   438: 'Spare_Fault_438', class No Acknowledgement, trigger "DB302_HMI_Faults_Carrier6_Faults_3" bit 5
   439: 'Spare_Fault_439', class No Acknowledgement, trigger "DB302_HMI_Faults_Carrier6_Faults_3" bit 6
   440: 'Spare_Fault_440', class No Acknowledgement, trigger "DB302_HMI_Faults_Carrier6_Faults_3" bit 7
   441: 'Spare_Fault_441', class No Acknowledgement, trigger "DB302_HMI_Faults_Carrier6_Faults_3" bit 8
   442: 'Spare_Fault_442', class No Acknowledgement, trigger "DB302_HMI_Faults_Carrier6_Faults_3" bit 9
   443: 'Spare_Fault_443', class No Acknowledgement, trigger "DB302_HMI_Faults_Carrier6_Faults_3" bit 10
   444: 'Spare_Fault_444', class No Acknowledgement, trigger "DB302_HMI_Faults_Carrier6_Faults_3" bit 11
   445: 'Spare_Fault_445', class No Acknowledgement, trigger "DB302_HMI_Faults_Carrier6_Faults_3" bit 12
   446: 'Spare_Fault_446', class No Acknowledgement, trigger "DB302_HMI_Faults_Carrier6_Faults_3" bit 13
   447: 'Spare_Fault_447', class No Acknowledgement, trigger "DB302_HMI_Faults_Carrier6_Faults_3" bit 14
   448: 'Spare_Fault_448', class No Acknowledgement, trigger "DB302_HMI_Faults_Carrier6_Faults_3" bit 15
   449: 'Carrier 07 Disconnect Open Power Fault DI11.0', class No Acknowledgement, trigger "DB302_HMI_Faults_Carrier7_Faults_0" bit 0
   450: 'Carrier 07 Drive Profinet Comm Fault', class No Acknowledgement, trigger "DB302_HMI_Faults_Carrier7_Faults_0" bit 1
   451: 'Carrier 07 Production Stop Not Reset', class No Acknowledgement, trigger "DB302_HMI_Faults_Carrier7_Faults_0" bit 2
   452: 'Carrier 07 CB02122 Tripped', class No Acknowledgement, trigger "DB302_HMI_Faults_Carrier7_Faults_0" bit 3
   453: 'Carrier 07 CB02123 Tripped', class No Acknowledgement, trigger "DB302_HMI_Faults_Carrier7_Faults_0" bit 4
   454: 'Carrier 07 AUX1 CB Tripped', class No Acknowledgement, trigger "DB302_HMI_Faults_Carrier7_Faults_0" bit 5
   455: 'Carrier 07 AUX2 CB Tripped', class No Acknowledgement, trigger "DB302_HMI_Faults_Carrier7_Faults_0" bit 6
   456: 'Carrier 07 PLC Not Communicating', class No Acknowledgement, trigger "DB302_HMI_Faults_Carrier7_Faults_0" bit 7
   457: 'Carrier 07 Safe Input Card Fault', class No Acknowledgement, trigger "DB302_HMI_Faults_Carrier7_Faults_0" bit 8
   458: 'Carrier 07 Safe Output Card Fault', class No Acknowledgement, trigger "DB302_HMI_Faults_Carrier7_Faults_0" bit 9
   459: 'Carrier 07 Standard Input Card Fault', class No Acknowledgement, trigger "DB302_HMI_Faults_Carrier7_Faults_0" bit 10
   460: 'Carrier 07 Standard Output Card Fault', class No Acknowledgement, trigger "DB302_HMI_Faults_Carrier7_Faults_0" bit 11
   461: 'Carrier 07 Encoder Position Fault', class No Acknowledgement, trigger "DB302_HMI_Faults_Carrier7_Faults_0" bit 12
   462: 'Carrier 07 Encoder Internal Error', class No Acknowledgement, trigger "DB302_HMI_Faults_Carrier7_Faults_0" bit 13
   463: 'Carrier 07 Encoder Comm Fault', class No Acknowledgement, trigger "DB302_HMI_Faults_Carrier7_Faults_0" bit 14
   464: 'Carrier 07 HMI Comm Fault', class No Acknowledgement, trigger "DB302_HMI_Faults_Carrier7_Faults_0" bit 15
   465: 'Carrier 07 Crash Detection Fault', class No Acknowledgement, trigger "DB302_HMI_Faults_Carrier7_Faults_1" bit 0
   466: 'Carrier 07 Carrier Number Invalid', class No Acknowledgement, trigger "DB302_HMI_Faults_Carrier7_Faults_1" bit 1
   467: 'Carrier 07 Drive: PROFINET configuration error', class No Acknowledgement, trigger "DB302_HMI_Faults_Carrier7_Faults_1" bit 2
   468: 'Carrier 07 Drive: Error internal communications', class No Acknowledgement, trigger "DB302_HMI_Faults_Carrier7_Faults_1" bit 3
   469: 'Carrier 07 Drive: Motor overtemperature', class No Acknowledgement, trigger "DB302_HMI_Faults_Carrier7_Faults_1" bit 4
   470: 'Carrier 07 Drive: Motor overcurrent', class No Acknowledgement, trigger "DB302_HMI_Faults_Carrier7_Faults_1" bit 5
   471: 'Carrier 07 Drive: Infeed or power unit not ready', class No Acknowledgement, trigger "DB302_HMI_Faults_Carrier7_Faults_1" bit 6
   472: 'Carrier 07 Drive: Short-circuit/ground fault detected', class No Acknowledgement, trigger "DB302_HMI_Faults_Carrier7_Faults_1" bit 7
   473: 'Carrier 07 Drive: PROFINET Setpoint timeout', class No Acknowledgement, trigger "DB302_HMI_Faults_Carrier7_Faults_1" bit 8
   474: 'Carrier 07 Power unit: Overcurrent', class No Acknowledgement, trigger "DB302_HMI_Faults_Carrier7_Faults_1" bit 9
   475: 'Carrier 07 Power unit: DC link voltage overvoltage', class No Acknowledgement, trigger "DB302_HMI_Faults_Carrier7_Faults_1" bit 10
   476: 'Carrier 07 Power unit: DC link voltage undervoltage', class No Acknowledgement, trigger "DB302_HMI_Faults_Carrier7_Faults_1" bit 11
   477: 'Carrier 07 Power unit: Line phase failure in main circuit', class No Acknowledgement, trigger "DB302_HMI_Faults_Carrier7_Faults_1" bit 12
   478: 'Carrier 07 Power unit: Phase failure motor cable', class No Acknowledgement, trigger "DB302_HMI_Faults_Carrier7_Faults_1" bit 13
   479: 'Carrier 07 Power unit: Ground fault', class No Acknowledgement, trigger "DB302_HMI_Faults_Carrier7_Faults_1" bit 14
   480: 'Spare_Fault_480', class No Acknowledgement, trigger "DB302_HMI_Faults_Carrier7_Faults_1" bit 15
   481: 'Carrier 07 Motion Off Fault', class No Acknowledgement, trigger "DB302_HMI_Faults_Carrier7_Faults_2" bit 0
   482: 'Carrier 07 Motion On Fault', class No Acknowledgement, trigger "DB302_HMI_Faults_Carrier7_Faults_2" bit 1
   483: 'Carrier 07 Spacing Fault', class No Acknowledgement, trigger "DB302_HMI_Faults_Carrier7_Faults_2" bit 2
   484: 'Carrier 07 Duplicate Carrier Number Fault', class No Acknowledgement, trigger "DB302_HMI_Faults_Carrier7_Faults_2" bit 3
   485: 'Spare_Fault_485', class No Acknowledgement, trigger "DB302_HMI_Faults_Carrier7_Faults_2" bit 4
   486: 'Spare_Fault_486', class No Acknowledgement, trigger "DB302_HMI_Faults_Carrier7_Faults_2" bit 5
   487: 'Spare_Fault_487', class No Acknowledgement, trigger "DB302_HMI_Faults_Carrier7_Faults_2" bit 6
   488: 'Spare_Fault_488', class No Acknowledgement, trigger "DB302_HMI_Faults_Carrier7_Faults_2" bit 7
   489: 'Spare_Fault_489', class No Acknowledgement, trigger "DB302_HMI_Faults_Carrier7_Faults_2" bit 8
   490: 'Spare_Fault_490', class No Acknowledgement, trigger "DB302_HMI_Faults_Carrier7_Faults_2" bit 9
   491: 'Spare_Fault_491', class No Acknowledgement, trigger "DB302_HMI_Faults_Carrier7_Faults_2" bit 10
   492: 'Spare_Fault_492', class No Acknowledgement, trigger "DB302_HMI_Faults_Carrier7_Faults_2" bit 11
   493: 'Spare_Fault_493', class No Acknowledgement, trigger "DB302_HMI_Faults_Carrier7_Faults_2" bit 12
   494: 'Spare_Fault_494', class No Acknowledgement, trigger "DB302_HMI_Faults_Carrier7_Faults_2" bit 13
   495: 'Spare_Fault_495', class No Acknowledgement, trigger "DB302_HMI_Faults_Carrier7_Faults_2" bit 14
   496: 'Spare_Fault_496', class No Acknowledgement, trigger "DB302_HMI_Faults_Carrier7_Faults_2" bit 15
   497: 'Spare_Fault_497', class No Acknowledgement, trigger "DB302_HMI_Faults_Carrier7_Faults_3" bit 0
   498: 'Spare_Fault_498', class No Acknowledgement, trigger "DB302_HMI_Faults_Carrier7_Faults_3" bit 1
   499: 'Spare_Fault_499', class No Acknowledgement, trigger "DB302_HMI_Faults_Carrier7_Faults_3" bit 2
   500: 'Spare_Fault_500', class No Acknowledgement, trigger "DB302_HMI_Faults_Carrier7_Faults_3" bit 3
   501: 'Spare_Fault_501', class No Acknowledgement, trigger "DB302_HMI_Faults_Carrier7_Faults_3" bit 4
   502: 'Spare_Fault_502', class No Acknowledgement, trigger "DB302_HMI_Faults_Carrier7_Faults_3" bit 5
   503: 'Spare_Fault_503', class No Acknowledgement, trigger "DB302_HMI_Faults_Carrier7_Faults_3" bit 6
   504: 'Spare_Fault_504', class No Acknowledgement, trigger "DB302_HMI_Faults_Carrier7_Faults_3" bit 7
   505: 'Spare_Fault_505', class No Acknowledgement, trigger "DB302_HMI_Faults_Carrier7_Faults_3" bit 8
   506: 'Spare_Fault_506', class No Acknowledgement, trigger "DB302_HMI_Faults_Carrier7_Faults_3" bit 9
   507: 'Spare_Fault_507', class No Acknowledgement, trigger "DB302_HMI_Faults_Carrier7_Faults_3" bit 10
   508: 'Spare_Fault_508', class No Acknowledgement, trigger "DB302_HMI_Faults_Carrier7_Faults_3" bit 11
   509: 'Spare_Fault_509', class No Acknowledgement, trigger "DB302_HMI_Faults_Carrier7_Faults_3" bit 12
   510: 'Spare_Fault_510', class No Acknowledgement, trigger "DB302_HMI_Faults_Carrier7_Faults_3" bit 13
   511: 'Spare_Fault_511', class No Acknowledgement, trigger "DB302_HMI_Faults_Carrier7_Faults_3" bit 14
   512: 'Spare_Fault_512', class No Acknowledgement, trigger "DB302_HMI_Faults_Carrier7_Faults_3" bit 15
   513: 'Carrier 08 Disconnect Open Power Fault DI11.0', class No Acknowledgement, trigger "DB302_HMI_Faults_Carrier8_Faults_0" bit 0
   514: 'Carrier 08 Drive Profinet Comm Fault', class No Acknowledgement, trigger "DB302_HMI_Faults_Carrier8_Faults_0" bit 1
   515: 'Carrier 08 Production Stop Not Reset', class No Acknowledgement, trigger "DB302_HMI_Faults_Carrier8_Faults_0" bit 2
   516: 'Carrier 08 CB02122 Tripped', class No Acknowledgement, trigger "DB302_HMI_Faults_Carrier8_Faults_0" bit 3
   517: 'Carrier 08 CB02123 Tripped', class No Acknowledgement, trigger "DB302_HMI_Faults_Carrier8_Faults_0" bit 4
   518: 'Carrier 08 AUX1 CB Tripped', class No Acknowledgement, trigger "DB302_HMI_Faults_Carrier8_Faults_0" bit 5
   519: 'Carrier 08 AUX2 CB Tripped', class No Acknowledgement, trigger "DB302_HMI_Faults_Carrier8_Faults_0" bit 6
   520: 'Carrier 08 PLC Not Communicating', class No Acknowledgement, trigger "DB302_HMI_Faults_Carrier8_Faults_0" bit 7
   521: 'Carrier 08 Safe Input Card Fault', class No Acknowledgement, trigger "DB302_HMI_Faults_Carrier8_Faults_0" bit 8
   522: 'Carrier 08 Safe Output Card Fault', class No Acknowledgement, trigger "DB302_HMI_Faults_Carrier8_Faults_0" bit 9
   523: 'Carrier 08 Standard Input Card Fault', class No Acknowledgement, trigger "DB302_HMI_Faults_Carrier8_Faults_0" bit 10
   524: 'Carrier 08 Standard Output Card Fault', class No Acknowledgement, trigger "DB302_HMI_Faults_Carrier8_Faults_0" bit 11
   525: 'Carrier 08 Encoder Position Fault', class No Acknowledgement, trigger "DB302_HMI_Faults_Carrier8_Faults_0" bit 12
   526: 'Carrier 08 Encoder Internal Error', class No Acknowledgement, trigger "DB302_HMI_Faults_Carrier8_Faults_0" bit 13
   527: 'Carrier 08 Encoder Comm Fault', class No Acknowledgement, trigger "DB302_HMI_Faults_Carrier8_Faults_0" bit 14
   528: 'Carrier 08 HMI Comm Fault', class No Acknowledgement, trigger "DB302_HMI_Faults_Carrier8_Faults_0" bit 15
   529: 'Carrier 08 Crash Detection Fault', class No Acknowledgement, trigger "DB302_HMI_Faults_Carrier8_Faults_1" bit 0
   530: 'Carrier 08 Carrier Number Invalid', class No Acknowledgement, trigger "DB302_HMI_Faults_Carrier8_Faults_1" bit 1
   531: 'Carrier 08 Drive: PROFINET configuration error', class No Acknowledgement, trigger "DB302_HMI_Faults_Carrier8_Faults_1" bit 2
   532: 'Carrier 08 Drive: Error internal communications', class No Acknowledgement, trigger "DB302_HMI_Faults_Carrier8_Faults_1" bit 3
   533: 'Carrier 08 Drive: Motor overtemperature', class No Acknowledgement, trigger "DB302_HMI_Faults_Carrier8_Faults_1" bit 4
   534: 'Carrier 08 Drive: Motor overcurrent', class No Acknowledgement, trigger "DB302_HMI_Faults_Carrier8_Faults_1" bit 5
   535: 'Carrier 08 Drive: Infeed or power unit not ready', class No Acknowledgement, trigger "DB302_HMI_Faults_Carrier8_Faults_1" bit 6
   536: 'Carrier 08 Drive: Short-circuit/ground fault detected', class No Acknowledgement, trigger "DB302_HMI_Faults_Carrier8_Faults_1" bit 7
   537: 'Carrier 08 Drive: PROFINET Setpoint timeout', class No Acknowledgement, trigger "DB302_HMI_Faults_Carrier8_Faults_1" bit 8
   538: 'Carrier 08 Power unit: Overcurrent', class No Acknowledgement, trigger "DB302_HMI_Faults_Carrier8_Faults_1" bit 9
   539: 'Carrier 08 Power unit: DC link voltage overvoltage', class No Acknowledgement, trigger "DB302_HMI_Faults_Carrier8_Faults_1" bit 10
   540: 'Carrier 08 Power unit: DC link voltage undervoltage', class No Acknowledgement, trigger "DB302_HMI_Faults_Carrier8_Faults_1" bit 11
   541: 'Carrier 08 Power unit: Line phase failure in main circuit', class No Acknowledgement, trigger "DB302_HMI_Faults_Carrier8_Faults_1" bit 12
   542: 'Carrier 08 Power unit: Phase failure motor cable', class No Acknowledgement, trigger "DB302_HMI_Faults_Carrier8_Faults_1" bit 13
   543: 'Carrier 08 Power unit: Ground fault', class No Acknowledgement, trigger "DB302_HMI_Faults_Carrier8_Faults_1" bit 14
   544: 'Spare_Fault_544', class No Acknowledgement, trigger "DB302_HMI_Faults_Carrier8_Faults_1" bit 15
   545: 'Carrier 08 Motion Off Fault', class No Acknowledgement, trigger "DB302_HMI_Faults_Carrier8_Faults_2" bit 0
   546: 'Carrier 08 Motion On Fault', class No Acknowledgement, trigger "DB302_HMI_Faults_Carrier8_Faults_2" bit 1
   547: 'Carrier 08 Spacing Fault', class No Acknowledgement, trigger "DB302_HMI_Faults_Carrier8_Faults_2" bit 2
   548: 'Carrier 08 Duplicate Carrier Number Fault', class No Acknowledgement, trigger "DB302_HMI_Faults_Carrier8_Faults_2" bit 3
   549: 'Spare_Fault_549', class No Acknowledgement, trigger "DB302_HMI_Faults_Carrier8_Faults_2" bit 4
   550: 'Spare_Fault_550', class No Acknowledgement, trigger "DB302_HMI_Faults_Carrier8_Faults_2" bit 5
   551: 'Spare_Fault_551', class No Acknowledgement, trigger "DB302_HMI_Faults_Carrier8_Faults_2" bit 6
   552: 'Spare_Fault_552', class No Acknowledgement, trigger "DB302_HMI_Faults_Carrier8_Faults_2" bit 7
   553: 'Spare_Fault_553', class No Acknowledgement, trigger "DB302_HMI_Faults_Carrier8_Faults_2" bit 8
   554: 'Spare_Fault_554', class No Acknowledgement, trigger "DB302_HMI_Faults_Carrier8_Faults_2" bit 9
   555: 'Spare_Fault_555', class No Acknowledgement, trigger "DB302_HMI_Faults_Carrier8_Faults_2" bit 10
   556: 'Spare_Fault_556', class No Acknowledgement, trigger "DB302_HMI_Faults_Carrier8_Faults_2" bit 11
   557: 'Spare_Fault_557', class No Acknowledgement, trigger "DB302_HMI_Faults_Carrier8_Faults_2" bit 12
   558: 'Spare_Fault_558', class No Acknowledgement, trigger "DB302_HMI_Faults_Carrier8_Faults_2" bit 13
   559: 'Spare_Fault_559', class No Acknowledgement, trigger "DB302_HMI_Faults_Carrier8_Faults_2" bit 14
   560: 'Spare_Fault_560', class No Acknowledgement, trigger "DB302_HMI_Faults_Carrier8_Faults_2" bit 15
   561: 'Spare_Fault_561', class No Acknowledgement, trigger "DB302_HMI_Faults_Carrier8_Faults_3" bit 0
   562: 'Spare_Fault_562', class No Acknowledgement, trigger "DB302_HMI_Faults_Carrier8_Faults_3" bit 1
   563: 'Spare_Fault_563', class No Acknowledgement, trigger "DB302_HMI_Faults_Carrier8_Faults_3" bit 2
   564: 'Spare_Fault_564', class No Acknowledgement, trigger "DB302_HMI_Faults_Carrier8_Faults_3" bit 3
   565: 'Spare_Fault_565', class No Acknowledgement, trigger "DB302_HMI_Faults_Carrier8_Faults_3" bit 4
   566: 'Spare_Fault_566', class No Acknowledgement, trigger "DB302_HMI_Faults_Carrier8_Faults_3" bit 5
   567: 'Spare_Fault_567', class No Acknowledgement, trigger "DB302_HMI_Faults_Carrier8_Faults_3" bit 6
   568: 'Spare_Fault_568', class No Acknowledgement, trigger "DB302_HMI_Faults_Carrier8_Faults_3" bit 7
   569: 'Spare_Fault_569', class No Acknowledgement, trigger "DB302_HMI_Faults_Carrier8_Faults_3" bit 8
   570: 'Spare_Fault_570', class No Acknowledgement, trigger "DB302_HMI_Faults_Carrier8_Faults_3" bit 9
   571: 'Spare_Fault_571', class No Acknowledgement, trigger "DB302_HMI_Faults_Carrier8_Faults_3" bit 10
   572: 'Spare_Fault_572', class No Acknowledgement, trigger "DB302_HMI_Faults_Carrier8_Faults_3" bit 11
   573: 'Spare_Fault_573', class No Acknowledgement, trigger "DB302_HMI_Faults_Carrier8_Faults_3" bit 12
   574: 'Spare_Fault_574', class No Acknowledgement, trigger "DB302_HMI_Faults_Carrier8_Faults_3" bit 13
   575: 'Spare_Fault_575', class No Acknowledgement, trigger "DB302_HMI_Faults_Carrier8_Faults_3" bit 14
   576: 'Spare_Fault_576', class No Acknowledgement, trigger "DB302_HMI_Faults_Carrier8_Faults_3" bit 15
   577: 'Carrier 09 Disconnect Open Power Fault DI11.0', class No Acknowledgement, trigger "DB302_HMI_Faults_Carrier9_Faults_0" bit 0
   578: 'Carrier 09 Drive Profinet Comm Fault', class No Acknowledgement, trigger "DB302_HMI_Faults_Carrier9_Faults_0" bit 1
   579: 'Carrier 09 Production Stop Not Reset', class No Acknowledgement, trigger "DB302_HMI_Faults_Carrier9_Faults_0" bit 2
   580: 'Carrier 09 CB02122 Tripped', class No Acknowledgement, trigger "DB302_HMI_Faults_Carrier9_Faults_0" bit 3
   581: 'Carrier 09 CB02123 Tripped', class No Acknowledgement, trigger "DB302_HMI_Faults_Carrier9_Faults_0" bit 4
   582: 'Carrier 09 AUX1 CB Tripped', class No Acknowledgement, trigger "DB302_HMI_Faults_Carrier9_Faults_0" bit 5
   583: 'Carrier 09 AUX2 CB Tripped', class No Acknowledgement, trigger "DB302_HMI_Faults_Carrier9_Faults_0" bit 6
   584: 'Carrier 09 PLC Not Communicating', class No Acknowledgement, trigger "DB302_HMI_Faults_Carrier9_Faults_0" bit 7
   585: 'Carrier 09 Safe Input Card Fault', class No Acknowledgement, trigger "DB302_HMI_Faults_Carrier9_Faults_0" bit 8
   586: 'Carrier 09 Safe Output Card Fault', class No Acknowledgement, trigger "DB302_HMI_Faults_Carrier9_Faults_0" bit 9
   587: 'Carrier 09 Standard Input Card Fault', class No Acknowledgement, trigger "DB302_HMI_Faults_Carrier9_Faults_0" bit 10
   588: 'Carrier 09 Standard Output Card Fault', class No Acknowledgement, trigger "DB302_HMI_Faults_Carrier9_Faults_0" bit 11
   589: 'Carrier 09 Encoder Position Fault', class No Acknowledgement, trigger "DB302_HMI_Faults_Carrier9_Faults_0" bit 12
   590: 'Carrier 09 Encoder Internal Error', class No Acknowledgement, trigger "DB302_HMI_Faults_Carrier9_Faults_0" bit 13
   591: 'Carrier 09 Encoder Comm Fault', class No Acknowledgement, trigger "DB302_HMI_Faults_Carrier9_Faults_0" bit 14
   592: 'Carrier 09 HMI Comm Fault', class No Acknowledgement, trigger "DB302_HMI_Faults_Carrier9_Faults_0" bit 15
   593: 'Carrier 09 Crash Detection Fault', class No Acknowledgement, trigger "DB302_HMI_Faults_Carrier9_Faults_1" bit 0
   594: 'Carrier 09 Carrier Number Invalid', class No Acknowledgement, trigger "DB302_HMI_Faults_Carrier9_Faults_1" bit 1
   595: 'Carrier 09 Drive: PROFINET configuration error', class No Acknowledgement, trigger "DB302_HMI_Faults_Carrier9_Faults_1" bit 2
   596: 'Carrier 09 Drive: Error internal communications', class No Acknowledgement, trigger "DB302_HMI_Faults_Carrier9_Faults_1" bit 3
   597: 'Carrier 09 Drive: Motor overtemperature', class No Acknowledgement, trigger "DB302_HMI_Faults_Carrier9_Faults_1" bit 4
   598: 'Carrier 09 Drive: Motor overcurrent', class No Acknowledgement, trigger "DB302_HMI_Faults_Carrier9_Faults_1" bit 5
   599: 'Carrier 09 Drive: Infeed or power unit not ready', class No Acknowledgement, trigger "DB302_HMI_Faults_Carrier9_Faults_1" bit 6
   600: 'Carrier 09 Drive: Short-circuit/ground fault detected', class No Acknowledgement, trigger "DB302_HMI_Faults_Carrier9_Faults_1" bit 7
   601: 'Carrier 09 Drive: PROFINET Setpoint timeout', class No Acknowledgement, trigger "DB302_HMI_Faults_Carrier9_Faults_1" bit 8
   602: 'Carrier 09 Power unit: Overcurrent', class No Acknowledgement, trigger "DB302_HMI_Faults_Carrier9_Faults_1" bit 9
   603: 'Carrier 09 Power unit: DC link voltage overvoltage', class No Acknowledgement, trigger "DB302_HMI_Faults_Carrier9_Faults_1" bit 10
   604: 'Carrier 09 Power unit: DC link voltage undervoltage', class No Acknowledgement, trigger "DB302_HMI_Faults_Carrier9_Faults_1" bit 11
   605: 'Carrier 09 Power unit: Line phase failure in main circuit', class No Acknowledgement, trigger "DB302_HMI_Faults_Carrier9_Faults_1" bit 12
   606: 'Carrier 09 Power unit: Phase failure motor cable', class No Acknowledgement, trigger "DB302_HMI_Faults_Carrier9_Faults_1" bit 13
   607: 'Carrier 09 Power unit: Ground fault', class No Acknowledgement, trigger "DB302_HMI_Faults_Carrier9_Faults_1" bit 14
   608: 'Spare_Fault_608', class No Acknowledgement, trigger "DB302_HMI_Faults_Carrier9_Faults_1" bit 15
   609: 'Carrier 09 Motion Off Fault', class No Acknowledgement, trigger "DB302_HMI_Faults_Carrier9_Faults_2" bit 0
   610: 'Carrier 09 Motion On Fault', class No Acknowledgement, trigger "DB302_HMI_Faults_Carrier9_Faults_2" bit 1
   611: 'Carrier 09 Spacing Fault', class No Acknowledgement, trigger "DB302_HMI_Faults_Carrier9_Faults_2" bit 2
   612: 'Carrier 09 Duplicate Carrier Number Fault', class No Acknowledgement, trigger "DB302_HMI_Faults_Carrier9_Faults_2" bit 3
   613: 'Spare_Fault_613', class No Acknowledgement, trigger "DB302_HMI_Faults_Carrier9_Faults_2" bit 4
   614: 'Spare_Fault_614', class No Acknowledgement, trigger "DB302_HMI_Faults_Carrier9_Faults_2" bit 5
   615: 'Spare_Fault_615', class No Acknowledgement, trigger "DB302_HMI_Faults_Carrier9_Faults_2" bit 6
   616: 'Spare_Fault_616', class No Acknowledgement, trigger "DB302_HMI_Faults_Carrier9_Faults_2" bit 7
   617: 'Spare_Fault_617', class No Acknowledgement, trigger "DB302_HMI_Faults_Carrier9_Faults_2" bit 8
   618: 'Spare_Fault_618', class No Acknowledgement, trigger "DB302_HMI_Faults_Carrier9_Faults_2" bit 9
   619: 'Spare_Fault_619', class No Acknowledgement, trigger "DB302_HMI_Faults_Carrier9_Faults_2" bit 10
   620: 'Spare_Fault_620', class No Acknowledgement, trigger "DB302_HMI_Faults_Carrier9_Faults_2" bit 11
   621: 'Spare_Fault_621', class No Acknowledgement, trigger "DB302_HMI_Faults_Carrier9_Faults_2" bit 12
   622: 'Spare_Fault_622', class No Acknowledgement, trigger "DB302_HMI_Faults_Carrier9_Faults_2" bit 13
   623: 'Spare_Fault_623', class No Acknowledgement, trigger "DB302_HMI_Faults_Carrier9_Faults_2" bit 14
   624: 'Spare_Fault_624', class No Acknowledgement, trigger "DB302_HMI_Faults_Carrier9_Faults_2" bit 15
   625: 'Spare_Fault_625', class No Acknowledgement, trigger "DB302_HMI_Faults_Carrier9_Faults_3" bit 0
   626: 'Spare_Fault_626', class No Acknowledgement, trigger "DB302_HMI_Faults_Carrier9_Faults_3" bit 1
   627: 'Spare_Fault_627', class No Acknowledgement, trigger "DB302_HMI_Faults_Carrier9_Faults_3" bit 2
   628: 'Spare_Fault_628', class No Acknowledgement, trigger "DB302_HMI_Faults_Carrier9_Faults_3" bit 3
   629: 'Spare_Fault_629', class No Acknowledgement, trigger "DB302_HMI_Faults_Carrier9_Faults_3" bit 4
   630: 'Spare_Fault_630', class No Acknowledgement, trigger "DB302_HMI_Faults_Carrier9_Faults_3" bit 5
   631: 'Spare_Fault_631', class No Acknowledgement, trigger "DB302_HMI_Faults_Carrier9_Faults_3" bit 6
   632: 'Spare_Fault_632', class No Acknowledgement, trigger "DB302_HMI_Faults_Carrier9_Faults_3" bit 7
   633: 'Spare_Fault_633', class No Acknowledgement, trigger "DB302_HMI_Faults_Carrier9_Faults_3" bit 8
   634: 'Spare_Fault_634', class No Acknowledgement, trigger "DB302_HMI_Faults_Carrier9_Faults_3" bit 9
   635: 'Spare_Fault_635', class No Acknowledgement, trigger "DB302_HMI_Faults_Carrier9_Faults_3" bit 10
   636: 'Spare_Fault_636', class No Acknowledgement, trigger "DB302_HMI_Faults_Carrier9_Faults_3" bit 11
   637: 'Spare_Fault_637', class No Acknowledgement, trigger "DB302_HMI_Faults_Carrier9_Faults_3" bit 12
   638: 'Spare_Fault_638', class No Acknowledgement, trigger "DB302_HMI_Faults_Carrier9_Faults_3" bit 13
   639: 'Spare_Fault_639', class No Acknowledgement, trigger "DB302_HMI_Faults_Carrier9_Faults_3" bit 14
   640: 'Spare_Fault_640', class No Acknowledgement, trigger "DB302_HMI_Faults_Carrier9_Faults_3" bit 15
   641: 'Carrier 10 Disconnect Open Power Fault DI11.0', class No Acknowledgement, trigger "DB302_HMI_Faults_Carrier10_Faults_0" bit 0
   642: 'Carrier 10 Drive Profinet Comm Fault', class No Acknowledgement, trigger "DB302_HMI_Faults_Carrier10_Faults_0" bit 1
   643: 'Carrier 10 Production Stop Not Reset', class No Acknowledgement, trigger "DB302_HMI_Faults_Carrier10_Faults_0" bit 2
   644: 'Carrier 10 CB02122 Tripped', class No Acknowledgement, trigger "DB302_HMI_Faults_Carrier10_Faults_0" bit 3
   645: 'Carrier 10 CB02123 Tripped', class No Acknowledgement, trigger "DB302_HMI_Faults_Carrier10_Faults_0" bit 4
   646: 'Carrier 10 AUX1 CB Tripped', class No Acknowledgement, trigger "DB302_HMI_Faults_Carrier10_Faults_0" bit 5
   647: 'Carrier 10 AUX2 CB Tripped', class No Acknowledgement, trigger "DB302_HMI_Faults_Carrier10_Faults_0" bit 6
   648: 'Carrier 10 PLC Not Communicating', class No Acknowledgement, trigger "DB302_HMI_Faults_Carrier10_Faults_0" bit 7
   649: 'Carrier 10 Safe Input Card Fault', class No Acknowledgement, trigger "DB302_HMI_Faults_Carrier10_Faults_0" bit 8
   650: 'Carrier 10 Safe Output Card Fault', class No Acknowledgement, trigger "DB302_HMI_Faults_Carrier10_Faults_0" bit 9
   651: 'Carrier 10 Standard Input Card Fault', class No Acknowledgement, trigger "DB302_HMI_Faults_Carrier10_Faults_0" bit 10
   652: 'Carrier 10 Standard Output Card Fault', class No Acknowledgement, trigger "DB302_HMI_Faults_Carrier10_Faults_0" bit 11
   653: 'Carrier 10 Encoder Position Fault', class No Acknowledgement, trigger "DB302_HMI_Faults_Carrier10_Faults_0" bit 12
   654: 'Carrier 10 Encoder Internal Error', class No Acknowledgement, trigger "DB302_HMI_Faults_Carrier10_Faults_0" bit 13
   655: 'Carrier 10 Encoder Comm Fault', class No Acknowledgement, trigger "DB302_HMI_Faults_Carrier10_Faults_0" bit 14
   656: 'Carrier 10 HMI Comm Fault', class No Acknowledgement, trigger "DB302_HMI_Faults_Carrier10_Faults_0" bit 15
   657: 'Carrier 10 Crash Detection Fault', class No Acknowledgement, trigger "DB302_HMI_Faults_Carrier10_Faults_1" bit 0
   658: 'Carrier 10 Carrier Number Invalid', class No Acknowledgement, trigger "DB302_HMI_Faults_Carrier10_Faults_1" bit 1
   659: 'Carrier 10 Drive: PROFINET configuration error', class No Acknowledgement, trigger "DB302_HMI_Faults_Carrier10_Faults_1" bit 2
   660: 'Carrier 10 Drive: Error internal communications', class No Acknowledgement, trigger "DB302_HMI_Faults_Carrier10_Faults_1" bit 3
   661: 'Carrier 10 Drive: Motor overtemperature', class No Acknowledgement, trigger "DB302_HMI_Faults_Carrier10_Faults_1" bit 4
   662: 'Carrier 10 Drive: Motor overcurrent', class No Acknowledgement, trigger "DB302_HMI_Faults_Carrier10_Faults_1" bit 5
   663: 'Carrier 10 Drive: Infeed or power unit not ready', class No Acknowledgement, trigger "DB302_HMI_Faults_Carrier10_Faults_1" bit 6
   664: 'Carrier 10 Drive: Short-circuit/ground fault detected', class No Acknowledgement, trigger "DB302_HMI_Faults_Carrier10_Faults_1" bit 7
   665: 'Carrier 10 Drive: PROFINET Setpoint timeout', class No Acknowledgement, trigger "DB302_HMI_Faults_Carrier10_Faults_1" bit 8
   666: 'Carrier 10 Power unit: Overcurrent', class No Acknowledgement, trigger "DB302_HMI_Faults_Carrier10_Faults_1" bit 9
   667: 'Carrier 10 Power unit: DC link voltage overvoltage', class No Acknowledgement, trigger "DB302_HMI_Faults_Carrier10_Faults_1" bit 10
   668: 'Carrier 10 Power unit: DC link voltage undervoltage', class No Acknowledgement, trigger "DB302_HMI_Faults_Carrier10_Faults_1" bit 11
   669: 'Carrier 10 Power unit: Line phase failure in main circuit', class No Acknowledgement, trigger "DB302_HMI_Faults_Carrier10_Faults_1" bit 12
   670: 'Carrier 10 Power unit: Phase failure motor cable', class No Acknowledgement, trigger "DB302_HMI_Faults_Carrier10_Faults_1" bit 13
   671: 'Carrier 10 Power unit: Ground fault', class No Acknowledgement, trigger "DB302_HMI_Faults_Carrier10_Faults_1" bit 14
   672: 'Spare_Fault_672', class No Acknowledgement, trigger "DB302_HMI_Faults_Carrier10_Faults_1" bit 15
   673: 'Carrier 10 Motion Off Fault', class No Acknowledgement, trigger "DB302_HMI_Faults_Carrier10_Faults_2" bit 0
   674: 'Carrier 10 Motion On Fault', class No Acknowledgement, trigger "DB302_HMI_Faults_Carrier10_Faults_2" bit 1
   675: 'Carrier 10 Spacing Fault', class No Acknowledgement, trigger "DB302_HMI_Faults_Carrier10_Faults_2" bit 2
   676: 'Carrier 10 Duplicate Carrier Number Fault', class No Acknowledgement, trigger "DB302_HMI_Faults_Carrier10_Faults_2" bit 3
   677: 'Spare_Fault_677', class No Acknowledgement, trigger "DB302_HMI_Faults_Carrier10_Faults_2" bit 4
   678: 'Spare_Fault_678', class No Acknowledgement, trigger "DB302_HMI_Faults_Carrier10_Faults_2" bit 5
   679: 'Spare_Fault_679', class No Acknowledgement, trigger "DB302_HMI_Faults_Carrier10_Faults_2" bit 6
   680: 'Spare_Fault_680', class No Acknowledgement, trigger "DB302_HMI_Faults_Carrier10_Faults_2" bit 7
   681: 'Spare_Fault_681', class No Acknowledgement, trigger "DB302_HMI_Faults_Carrier10_Faults_2" bit 8
   682: 'Spare_Fault_682', class No Acknowledgement, trigger "DB302_HMI_Faults_Carrier10_Faults_2" bit 9
   683: 'Spare_Fault_683', class No Acknowledgement, trigger "DB302_HMI_Faults_Carrier10_Faults_2" bit 10
   684: 'Spare_Fault_684', class No Acknowledgement, trigger "DB302_HMI_Faults_Carrier10_Faults_2" bit 11
   685: 'Spare_Fault_685', class No Acknowledgement, trigger "DB302_HMI_Faults_Carrier10_Faults_2" bit 12
   686: 'Spare_Fault_686', class No Acknowledgement, trigger "DB302_HMI_Faults_Carrier10_Faults_2" bit 13
   687: 'Spare_Fault_687', class No Acknowledgement, trigger "DB302_HMI_Faults_Carrier10_Faults_2" bit 14
   688: 'Spare_Fault_688', class No Acknowledgement, trigger "DB302_HMI_Faults_Carrier10_Faults_2" bit 15
   689: 'Spare_Fault_689', class No Acknowledgement, trigger "DB302_HMI_Faults_Carrier10_Faults_3" bit 0
   690: 'Spare_Fault_690', class No Acknowledgement, trigger "DB302_HMI_Faults_Carrier10_Faults_3" bit 1
   691: 'Spare_Fault_691', class No Acknowledgement, trigger "DB302_HMI_Faults_Carrier10_Faults_3" bit 2
   692: 'Spare_Fault_692', class No Acknowledgement, trigger "DB302_HMI_Faults_Carrier10_Faults_3" bit 3
   693: 'Spare_Fault_693', class No Acknowledgement, trigger "DB302_HMI_Faults_Carrier10_Faults_3" bit 4
   694: 'Spare_Fault_694', class No Acknowledgement, trigger "DB302_HMI_Faults_Carrier10_Faults_3" bit 5
   695: 'Spare_Fault_695', class No Acknowledgement, trigger "DB302_HMI_Faults_Carrier10_Faults_3" bit 6
   696: 'Spare_Fault_696', class No Acknowledgement, trigger "DB302_HMI_Faults_Carrier10_Faults_3" bit 7
   697: 'Spare_Fault_697', class No Acknowledgement, trigger "DB302_HMI_Faults_Carrier10_Faults_3" bit 8
   698: 'Spare_Fault_698', class No Acknowledgement, trigger "DB302_HMI_Faults_Carrier10_Faults_3" bit 9
   699: 'Spare_Fault_699', class No Acknowledgement, trigger "DB302_HMI_Faults_Carrier10_Faults_3" bit 10
   700: 'Spare_Fault_700', class No Acknowledgement, trigger "DB302_HMI_Faults_Carrier10_Faults_3" bit 11
   701: 'Spare_Fault_701', class No Acknowledgement, trigger "DB302_HMI_Faults_Carrier10_Faults_3" bit 12
   702: 'Spare_Fault_702', class No Acknowledgement, trigger "DB302_HMI_Faults_Carrier10_Faults_3" bit 13
   703: 'Spare_Fault_703', class No Acknowledgement, trigger "DB302_HMI_Faults_Carrier10_Faults_3" bit 14
   704: 'Spare_Fault_704', class No Acknowledgement, trigger "DB302_HMI_Faults_Carrier10_Faults_3" bit 15
   705: 'Carrier 11 Disconnect Open Power Fault DI11.0', class No Acknowledgement, trigger "DB302_HMI_Faults_Carrier11_Faults_0" bit 0
   706: 'Carrier 11 Drive Profinet Comm Fault', class No Acknowledgement, trigger "DB302_HMI_Faults_Carrier11_Faults_0" bit 1
   707: 'Carrier 11 Production Stop Not Reset', class No Acknowledgement, trigger "DB302_HMI_Faults_Carrier11_Faults_0" bit 2
   708: 'Carrier 11 CB02122 Tripped', class No Acknowledgement, trigger "DB302_HMI_Faults_Carrier11_Faults_0" bit 3
   709: 'Carrier 11 CB02123 Tripped', class No Acknowledgement, trigger "DB302_HMI_Faults_Carrier11_Faults_0" bit 4
   710: 'Carrier 11 AUX1 CB Tripped', class No Acknowledgement, trigger "DB302_HMI_Faults_Carrier11_Faults_0" bit 5
   711: 'Carrier 11 AUX2 CB Tripped', class No Acknowledgement, trigger "DB302_HMI_Faults_Carrier11_Faults_0" bit 6
   712: 'Carrier 11 PLC Not Communicating', class No Acknowledgement, trigger "DB302_HMI_Faults_Carrier11_Faults_0" bit 7
   713: 'Carrier 11 Safe Input Card Fault', class No Acknowledgement, trigger "DB302_HMI_Faults_Carrier11_Faults_0" bit 8
   714: 'Carrier 11 Safe Output Card Fault', class No Acknowledgement, trigger "DB302_HMI_Faults_Carrier11_Faults_0" bit 9
   715: 'Carrier 11 Standard Input Card Fault', class No Acknowledgement, trigger "DB302_HMI_Faults_Carrier11_Faults_0" bit 10
   716: 'Carrier 11 Standard Output Card Fault', class No Acknowledgement, trigger "DB302_HMI_Faults_Carrier11_Faults_0" bit 11
   717: 'Carrier 11 Encoder Position Fault', class No Acknowledgement, trigger "DB302_HMI_Faults_Carrier11_Faults_0" bit 12
   718: 'Carrier 11 Encoder Internal Error', class No Acknowledgement, trigger "DB302_HMI_Faults_Carrier11_Faults_0" bit 13
   719: 'Carrier 11 Encoder Comm Fault', class No Acknowledgement, trigger "DB302_HMI_Faults_Carrier11_Faults_0" bit 14
   720: 'Carrier 11 HMI Comm Fault', class No Acknowledgement, trigger "DB302_HMI_Faults_Carrier11_Faults_0" bit 15
   721: 'Carrier 11 Crash Detection Fault', class No Acknowledgement, trigger "DB302_HMI_Faults_Carrier11_Faults_1" bit 0
   722: 'Carrier 11 Carrier Number Invalid', class No Acknowledgement, trigger "DB302_HMI_Faults_Carrier11_Faults_1" bit 1
   723: 'Carrier 11 Drive: PROFINET configuration error', class No Acknowledgement, trigger "DB302_HMI_Faults_Carrier11_Faults_1" bit 2
   724: 'Carrier 11 Drive: Error internal communications', class No Acknowledgement, trigger "DB302_HMI_Faults_Carrier11_Faults_1" bit 3
   725: 'Carrier 11 Drive: Motor overtemperature', class No Acknowledgement, trigger "DB302_HMI_Faults_Carrier11_Faults_1" bit 4
   726: 'Carrier 11 Drive: Motor overcurrent', class No Acknowledgement, trigger "DB302_HMI_Faults_Carrier11_Faults_1" bit 5
   727: 'Carrier 11 Drive: Infeed or power unit not ready', class No Acknowledgement, trigger "DB302_HMI_Faults_Carrier11_Faults_1" bit 6
   728: 'Carrier 11 Drive: Short-circuit/ground fault detected', class No Acknowledgement, trigger "DB302_HMI_Faults_Carrier11_Faults_1" bit 7
   729: 'Carrier 11 Drive: PROFINET Setpoint timeout', class No Acknowledgement, trigger "DB302_HMI_Faults_Carrier11_Faults_1" bit 8
   730: 'Carrier 11 Power unit: Overcurrent', class No Acknowledgement, trigger "DB302_HMI_Faults_Carrier11_Faults_1" bit 9
   731: 'Carrier 11 Power unit: DC link voltage overvoltage', class No Acknowledgement, trigger "DB302_HMI_Faults_Carrier11_Faults_1" bit 10
   732: 'Carrier 11 Power unit: DC link voltage undervoltage', class No Acknowledgement, trigger "DB302_HMI_Faults_Carrier11_Faults_1" bit 11
   733: 'Carrier 11 Power unit: Line phase failure in main circuit', class No Acknowledgement, trigger "DB302_HMI_Faults_Carrier11_Faults_1" bit 12
   734: 'Carrier 11 Power unit: Phase failure motor cable', class No Acknowledgement, trigger "DB302_HMI_Faults_Carrier11_Faults_1" bit 13
   735: 'Carrier 11 Power unit: Ground fault', class No Acknowledgement, trigger "DB302_HMI_Faults_Carrier11_Faults_1" bit 14
   736: 'Spare_Fault_736', class No Acknowledgement, trigger "DB302_HMI_Faults_Carrier11_Faults_1" bit 15
   737: 'Carrier 11 Motion Off Fault', class No Acknowledgement, trigger "DB302_HMI_Faults_Carrier11_Faults_2" bit 0
   738: 'Carrier 11 Motion On Fault', class No Acknowledgement, trigger "DB302_HMI_Faults_Carrier11_Faults_2" bit 1
   739: 'Carrier 11 Spacing Fault', class No Acknowledgement, trigger "DB302_HMI_Faults_Carrier11_Faults_2" bit 2
   740: 'Carrier 11 Duplicate Carrier Number Fault', class No Acknowledgement, trigger "DB302_HMI_Faults_Carrier11_Faults_2" bit 3
   741: 'Spare_Fault_741', class No Acknowledgement, trigger "DB302_HMI_Faults_Carrier11_Faults_2" bit 4
   742: 'Spare_Fault_742', class No Acknowledgement, trigger "DB302_HMI_Faults_Carrier11_Faults_2" bit 5
   743: 'Spare_Fault_743', class No Acknowledgement, trigger "DB302_HMI_Faults_Carrier11_Faults_2" bit 6
   744: 'Spare_Fault_744', class No Acknowledgement, trigger "DB302_HMI_Faults_Carrier11_Faults_2" bit 7
   745: 'Spare_Fault_745', class No Acknowledgement, trigger "DB302_HMI_Faults_Carrier11_Faults_2" bit 8
   746: 'Spare_Fault_746', class No Acknowledgement, trigger "DB302_HMI_Faults_Carrier11_Faults_2" bit 9
   747: 'Spare_Fault_747', class No Acknowledgement, trigger "DB302_HMI_Faults_Carrier11_Faults_2" bit 10
   748: 'Spare_Fault_748', class No Acknowledgement, trigger "DB302_HMI_Faults_Carrier11_Faults_2" bit 11
   749: 'Spare_Fault_749', class No Acknowledgement, trigger "DB302_HMI_Faults_Carrier11_Faults_2" bit 12
   750: 'Spare_Fault_750', class No Acknowledgement, trigger "DB302_HMI_Faults_Carrier11_Faults_2" bit 13
   751: 'Spare_Fault_751', class No Acknowledgement, trigger "DB302_HMI_Faults_Carrier11_Faults_2" bit 14
   752: 'Spare_Fault_752', class No Acknowledgement, trigger "DB302_HMI_Faults_Carrier11_Faults_2" bit 15
   753: 'Spare_Fault_753', class No Acknowledgement, trigger "DB302_HMI_Faults_Carrier11_Faults_3" bit 0
   754: 'Spare_Fault_754', class No Acknowledgement, trigger "DB302_HMI_Faults_Carrier11_Faults_3" bit 1
   755: 'Spare_Fault_755', class No Acknowledgement, trigger "DB302_HMI_Faults_Carrier11_Faults_3" bit 2
   756: 'Spare_Fault_756', class No Acknowledgement, trigger "DB302_HMI_Faults_Carrier11_Faults_3" bit 3
   757: 'Spare_Fault_757', class No Acknowledgement, trigger "DB302_HMI_Faults_Carrier11_Faults_3" bit 4
   758: 'Spare_Fault_758', class No Acknowledgement, trigger "DB302_HMI_Faults_Carrier11_Faults_3" bit 5
   759: 'Spare_Fault_759', class No Acknowledgement, trigger "DB302_HMI_Faults_Carrier11_Faults_3" bit 6
   760: 'Spare_Fault_760', class No Acknowledgement, trigger "DB302_HMI_Faults_Carrier11_Faults_3" bit 7
   761: 'Spare_Fault_761', class No Acknowledgement, trigger "DB302_HMI_Faults_Carrier11_Faults_3" bit 8
   762: 'Spare_Fault_762', class No Acknowledgement, trigger "DB302_HMI_Faults_Carrier11_Faults_3" bit 9
   763: 'Spare_Fault_763', class No Acknowledgement, trigger "DB302_HMI_Faults_Carrier11_Faults_3" bit 10
   764: 'Spare_Fault_764', class No Acknowledgement, trigger "DB302_HMI_Faults_Carrier11_Faults_3" bit 11
   765: 'Spare_Fault_765', class No Acknowledgement, trigger "DB302_HMI_Faults_Carrier11_Faults_3" bit 12
   766: 'Spare_Fault_766', class No Acknowledgement, trigger "DB302_HMI_Faults_Carrier11_Faults_3" bit 13
   767: 'Spare_Fault_767', class No Acknowledgement, trigger "DB302_HMI_Faults_Carrier11_Faults_3" bit 14
   768: 'Spare_Fault_768', class No Acknowledgement, trigger "DB302_HMI_Faults_Carrier11_Faults_3" bit 15
   769: 'Carrier 12 Disconnect Open Power Fault DI11.0', class No Acknowledgement, trigger "DB302_HMI_Faults_Carrier12_Faults_0" bit 0
   770: 'Carrier 12 Drive Profinet Comm Fault', class No Acknowledgement, trigger "DB302_HMI_Faults_Carrier12_Faults_0" bit 1
   771: 'Carrier 12 Production Stop Not Reset', class No Acknowledgement, trigger "DB302_HMI_Faults_Carrier12_Faults_0" bit 2
   772: 'Carrier 12 CB02122 Tripped', class No Acknowledgement, trigger "DB302_HMI_Faults_Carrier12_Faults_0" bit 3
   773: 'Carrier 12 CB02123 Tripped', class No Acknowledgement, trigger "DB302_HMI_Faults_Carrier12_Faults_0" bit 4
   774: 'Carrier 12 AUX1 CB Tripped', class No Acknowledgement, trigger "DB302_HMI_Faults_Carrier12_Faults_0" bit 5
   775: 'Carrier 12 AUX2 CB Tripped', class No Acknowledgement, trigger "DB302_HMI_Faults_Carrier12_Faults_0" bit 6
   776: 'Carrier 12 PLC Not Communicating', class No Acknowledgement, trigger "DB302_HMI_Faults_Carrier12_Faults_0" bit 7
   777: 'Carrier 12 Safe Input Card Fault', class No Acknowledgement, trigger "DB302_HMI_Faults_Carrier12_Faults_0" bit 8
   778: 'Carrier 12 Safe Output Card Fault', class No Acknowledgement, trigger "DB302_HMI_Faults_Carrier12_Faults_0" bit 9
   779: 'Carrier 12 Standard Input Card Fault', class No Acknowledgement, trigger "DB302_HMI_Faults_Carrier12_Faults_0" bit 10
   780: 'Carrier 12 Standard Output Card Fault', class No Acknowledgement, trigger "DB302_HMI_Faults_Carrier12_Faults_0" bit 11
   781: 'Carrier 12 Encoder Position Fault', class No Acknowledgement, trigger "DB302_HMI_Faults_Carrier12_Faults_0" bit 12
   782: 'Carrier 12 Encoder Internal Error', class No Acknowledgement, trigger "DB302_HMI_Faults_Carrier12_Faults_0" bit 13
   783: 'Carrier 12 Encoder Comm Fault', class No Acknowledgement, trigger "DB302_HMI_Faults_Carrier12_Faults_0" bit 14
   784: 'Carrier 12 HMI Comm Fault', class No Acknowledgement, trigger "DB302_HMI_Faults_Carrier12_Faults_0" bit 15
   785: 'Carrier 12 Crash Detection Fault', class No Acknowledgement, trigger "DB302_HMI_Faults_Carrier12_Faults_1" bit 0
   786: 'Carrier 12 Carrier Number Invalid', class No Acknowledgement, trigger "DB302_HMI_Faults_Carrier12_Faults_1" bit 1
   787: 'Carrier 12 Drive: PROFINET configuration error', class No Acknowledgement, trigger "DB302_HMI_Faults_Carrier12_Faults_1" bit 2
   788: 'Carrier 12 Drive: Error internal communications', class No Acknowledgement, trigger "DB302_HMI_Faults_Carrier12_Faults_1" bit 3
   789: 'Carrier 12 Drive: Motor overtemperature', class No Acknowledgement, trigger "DB302_HMI_Faults_Carrier12_Faults_1" bit 4
   790: 'Carrier 12 Drive: Motor overcurrent', class No Acknowledgement, trigger "DB302_HMI_Faults_Carrier12_Faults_1" bit 5
   791: 'Carrier 12 Drive: Infeed or power unit not ready', class No Acknowledgement, trigger "DB302_HMI_Faults_Carrier12_Faults_1" bit 6
   792: 'Carrier 12 Drive: Short-circuit/ground fault detected', class No Acknowledgement, trigger "DB302_HMI_Faults_Carrier12_Faults_1" bit 7
   793: 'Carrier 12 Drive: PROFINET Setpoint timeout', class No Acknowledgement, trigger "DB302_HMI_Faults_Carrier12_Faults_1" bit 8
   794: 'Carrier 12 Power unit: Overcurrent', class No Acknowledgement, trigger "DB302_HMI_Faults_Carrier12_Faults_1" bit 9
   795: 'Carrier 12 Power unit: DC link voltage overvoltage', class No Acknowledgement, trigger "DB302_HMI_Faults_Carrier12_Faults_1" bit 10
   796: 'Carrier 12 Power unit: DC link voltage undervoltage', class No Acknowledgement, trigger "DB302_HMI_Faults_Carrier12_Faults_1" bit 11
   797: 'Carrier 12 Power unit: Line phase failure in main circuit', class No Acknowledgement, trigger "DB302_HMI_Faults_Carrier12_Faults_1" bit 12
   798: 'Carrier 12 Power unit: Phase failure motor cable', class No Acknowledgement, trigger "DB302_HMI_Faults_Carrier12_Faults_1" bit 13
   799: 'Carrier 12 Power unit: Ground fault', class No Acknowledgement, trigger "DB302_HMI_Faults_Carrier12_Faults_1" bit 14
   800: 'Spare_Fault_800', class No Acknowledgement, trigger "DB302_HMI_Faults_Carrier12_Faults_1" bit 15
   801: 'Carrier 12 Motion Off Fault', class No Acknowledgement, trigger "DB302_HMI_Faults_Carrier12_Faults_2" bit 0
   802: 'Carrier 12 Motion On Fault', class No Acknowledgement, trigger "DB302_HMI_Faults_Carrier12_Faults_2" bit 1
   803: 'Carrier 12 Spacing Fault', class No Acknowledgement, trigger "DB302_HMI_Faults_Carrier12_Faults_2" bit 2
   804: 'Carrier 12 Duplicate Carrier Number Fault', class No Acknowledgement, trigger "DB302_HMI_Faults_Carrier12_Faults_2" bit 3
   805: 'Spare_Fault_805', class No Acknowledgement, trigger "DB302_HMI_Faults_Carrier12_Faults_2" bit 4
   806: 'Spare_Fault_806', class No Acknowledgement, trigger "DB302_HMI_Faults_Carrier12_Faults_2" bit 5
   807: 'Spare_Fault_807', class No Acknowledgement, trigger "DB302_HMI_Faults_Carrier12_Faults_2" bit 6
   808: 'Spare_Fault_808', class No Acknowledgement, trigger "DB302_HMI_Faults_Carrier12_Faults_2" bit 7
   809: 'Spare_Fault_809', class No Acknowledgement, trigger "DB302_HMI_Faults_Carrier12_Faults_2" bit 8
   810: 'Spare_Fault_810', class No Acknowledgement, trigger "DB302_HMI_Faults_Carrier12_Faults_2" bit 9
   811: 'Spare_Fault_811', class No Acknowledgement, trigger "DB302_HMI_Faults_Carrier12_Faults_2" bit 10
   812: 'Spare_Fault_812', class No Acknowledgement, trigger "DB302_HMI_Faults_Carrier12_Faults_2" bit 11
   813: 'Spare_Fault_813', class No Acknowledgement, trigger "DB302_HMI_Faults_Carrier12_Faults_2" bit 12
   814: 'Spare_Fault_814', class No Acknowledgement, trigger "DB302_HMI_Faults_Carrier12_Faults_2" bit 13
   815: 'Spare_Fault_815', class No Acknowledgement, trigger "DB302_HMI_Faults_Carrier12_Faults_2" bit 14
   816: 'Spare_Fault_816', class No Acknowledgement, trigger "DB302_HMI_Faults_Carrier12_Faults_2" bit 15
   817: 'Spare_Fault_817', class No Acknowledgement, trigger "DB302_HMI_Faults_Carrier12_Faults_3" bit 0
   818: 'Spare_Fault_818', class No Acknowledgement, trigger "DB302_HMI_Faults_Carrier12_Faults_3" bit 1
   819: 'Spare_Fault_819', class No Acknowledgement, trigger "DB302_HMI_Faults_Carrier12_Faults_3" bit 2
   820: 'Spare_Fault_820', class No Acknowledgement, trigger "DB302_HMI_Faults_Carrier12_Faults_3" bit 3
   821: 'Spare_Fault_821', class No Acknowledgement, trigger "DB302_HMI_Faults_Carrier12_Faults_3" bit 4
   822: 'Spare_Fault_822', class No Acknowledgement, trigger "DB302_HMI_Faults_Carrier12_Faults_3" bit 5
   823: 'Spare_Fault_823', class No Acknowledgement, trigger "DB302_HMI_Faults_Carrier12_Faults_3" bit 6
   824: 'Spare_Fault_824', class No Acknowledgement, trigger "DB302_HMI_Faults_Carrier12_Faults_3" bit 7
   825: 'Spare_Fault_825', class No Acknowledgement, trigger "DB302_HMI_Faults_Carrier12_Faults_3" bit 8
   826: 'Spare_Fault_826', class No Acknowledgement, trigger "DB302_HMI_Faults_Carrier12_Faults_3" bit 9
   827: 'Spare_Fault_827', class No Acknowledgement, trigger "DB302_HMI_Faults_Carrier12_Faults_3" bit 10
   828: 'Spare_Fault_828', class No Acknowledgement, trigger "DB302_HMI_Faults_Carrier12_Faults_3" bit 11
   829: 'Spare_Fault_829', class No Acknowledgement, trigger "DB302_HMI_Faults_Carrier12_Faults_3" bit 12
   830: 'Spare_Fault_830', class No Acknowledgement, trigger "DB302_HMI_Faults_Carrier12_Faults_3" bit 13
   831: 'Spare_Fault_831', class No Acknowledgement, trigger "DB302_HMI_Faults_Carrier12_Faults_3" bit 14
   832: 'Spare_Fault_832', class No Acknowledgement, trigger "DB302_HMI_Faults_Carrier12_Faults_3" bit 15
   833: 'Carrier 13 Disconnect Open Power Fault DI11.0', class No Acknowledgement, trigger "DB302_HMI_Faults_Carrier13_Faults_0" bit 0
   834: 'Carrier 13 Drive Profinet Comm Fault', class No Acknowledgement, trigger "DB302_HMI_Faults_Carrier13_Faults_0" bit 1
   835: 'Carrier 13 Production Stop Not Reset', class No Acknowledgement, trigger "DB302_HMI_Faults_Carrier13_Faults_0" bit 2
   836: 'Carrier 13 CB02122 Tripped', class No Acknowledgement, trigger "DB302_HMI_Faults_Carrier13_Faults_0" bit 3
   837: 'Carrier 13 CB02123 Tripped', class No Acknowledgement, trigger "DB302_HMI_Faults_Carrier13_Faults_0" bit 4
   838: 'Carrier 13 AUX1 CB Tripped', class No Acknowledgement, trigger "DB302_HMI_Faults_Carrier13_Faults_0" bit 5
   839: 'Carrier 13 AUX2 CB Tripped', class No Acknowledgement, trigger "DB302_HMI_Faults_Carrier13_Faults_0" bit 6
   840: 'Carrier 13 PLC Not Communicating', class No Acknowledgement, trigger "DB302_HMI_Faults_Carrier13_Faults_0" bit 7
   841: 'Carrier 13 Safe Input Card Fault', class No Acknowledgement, trigger "DB302_HMI_Faults_Carrier13_Faults_0" bit 8
   842: 'Carrier 13 Safe Output Card Fault', class No Acknowledgement, trigger "DB302_HMI_Faults_Carrier13_Faults_0" bit 9
   843: 'Carrier 13 Standard Input Card Fault', class No Acknowledgement, trigger "DB302_HMI_Faults_Carrier13_Faults_0" bit 10
   844: 'Carrier 13 Standard Output Card Fault', class No Acknowledgement, trigger "DB302_HMI_Faults_Carrier13_Faults_0" bit 11
   845: 'Carrier 13 Encoder Position Fault', class No Acknowledgement, trigger "DB302_HMI_Faults_Carrier13_Faults_0" bit 12
   846: 'Carrier 13 Encoder Internal Error', class No Acknowledgement, trigger "DB302_HMI_Faults_Carrier13_Faults_0" bit 13
   847: 'Carrier 13 Encoder Comm Fault', class No Acknowledgement, trigger "DB302_HMI_Faults_Carrier13_Faults_0" bit 14
   848: 'Carrier 13 HMI Comm Fault', class No Acknowledgement, trigger "DB302_HMI_Faults_Carrier13_Faults_0" bit 15
   849: 'Carrier 13 Crash Detection Fault', class No Acknowledgement, trigger "DB302_HMI_Faults_Carrier13_Faults_1" bit 0
   850: 'Carrier 13 Carrier Number Invalid', class No Acknowledgement, trigger "DB302_HMI_Faults_Carrier13_Faults_1" bit 1
   851: 'Carrier 13 Drive: PROFINET configuration error', class No Acknowledgement, trigger "DB302_HMI_Faults_Carrier13_Faults_1" bit 2
   852: 'Carrier 13 Drive: Error internal communications', class No Acknowledgement, trigger "DB302_HMI_Faults_Carrier13_Faults_1" bit 3
   853: 'Carrier 13 Drive: Motor overtemperature', class No Acknowledgement, trigger "DB302_HMI_Faults_Carrier13_Faults_1" bit 4
   854: 'Carrier 13 Drive: Motor overcurrent', class No Acknowledgement, trigger "DB302_HMI_Faults_Carrier13_Faults_1" bit 5
   855: 'Carrier 13 Drive: Infeed or power unit not ready', class No Acknowledgement, trigger "DB302_HMI_Faults_Carrier13_Faults_1" bit 6
   856: 'Carrier 13 Drive: Short-circuit/ground fault detected', class No Acknowledgement, trigger "DB302_HMI_Faults_Carrier13_Faults_1" bit 7
   857: 'Carrier 13 Drive: PROFINET Setpoint timeout', class No Acknowledgement, trigger "DB302_HMI_Faults_Carrier13_Faults_1" bit 8
   858: 'Carrier 13 Power unit: Overcurrent', class No Acknowledgement, trigger "DB302_HMI_Faults_Carrier13_Faults_1" bit 9
   859: 'Carrier 13 Power unit: DC link voltage overvoltage', class No Acknowledgement, trigger "DB302_HMI_Faults_Carrier13_Faults_1" bit 10
   860: 'Carrier 13 Power unit: DC link voltage undervoltage', class No Acknowledgement, trigger "DB302_HMI_Faults_Carrier13_Faults_1" bit 11
   861: 'Carrier 13 Power unit: Line phase failure in main circuit', class No Acknowledgement, trigger "DB302_HMI_Faults_Carrier13_Faults_1" bit 12
   862: 'Carrier 13 Power unit: Phase failure motor cable', class No Acknowledgement, trigger "DB302_HMI_Faults_Carrier13_Faults_1" bit 13
   863: 'Carrier 13 Power unit: Ground fault', class No Acknowledgement, trigger "DB302_HMI_Faults_Carrier13_Faults_1" bit 14
